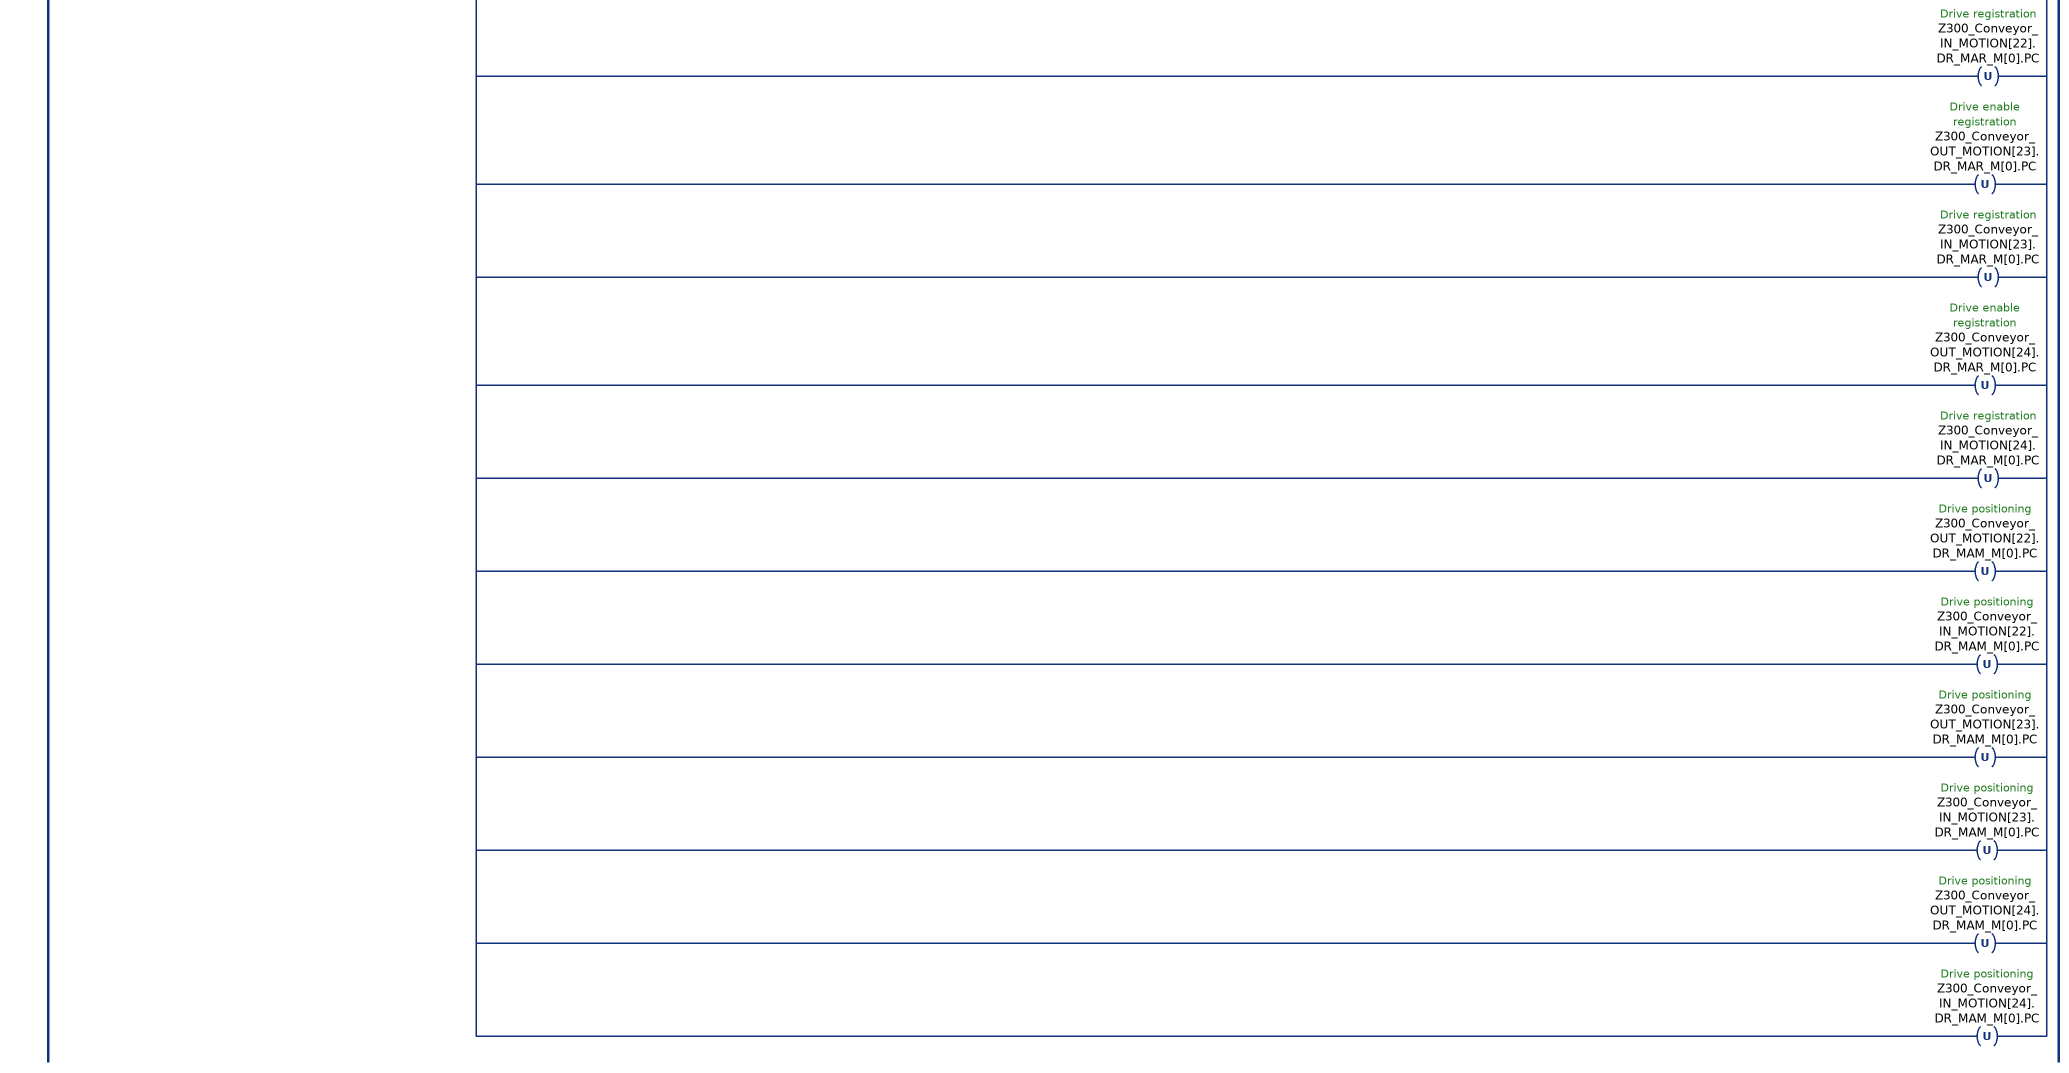
   // Positioning request (In case of head positioning also previous conveyors are involved)
   32: XIO(M310Popup[0].ST_xPlateInPositionToRise)XIO(M310Popup[1].ST_xPlateInPositionToRise)XIC(M310Popup[0].AUX_tSearchPlateData.xPlateHooked)[XIC(M310Popup[0].ST_xPlateToSinglePositioning) XIO(Z300_LineTracking.rgtTrkConv[22].xGlassPresence) XIO(Z300_LineTracking.rgtTrkConv[23].xGlassPresence) XIO(M310Popup[0].ST_xPlatePresence) [XIO(M310Popup[0].ST_xPlateUnderPopup) ,XIO(xDebugOFF) ] XIC(M310Popup[0].ST_xOutputEnable) XIC(M310Popup[0].INPUT_xPopupLow) XIC(M310Popup[0].ST_xInitialConditionForRise) ,XIC(M310Popup[1].ST_xPlateToSinglePositioning) XIO(Z300_LineTracking.rgtTrkConv[22].xGlassPresence) XIO(Z300_LineTracking.rgtTrkConv[23].xGlassPresence) XIO(Z300_LineTracking.rgtTrkConv[24].xGlassPresence) XIO(M310Popup[1].ST_xPlatePresence) XIO(M310Popup[0].ST_xPlateUnderPopup) [XIO(M310Popup[1].ST_xPlateUnderPopup) ,XIO(xDebugOFF) ] XIC(M310Popup[1].ST_xOutputEnable) XIC(M310Popup[1].INPUT_xPopupLow) XIC(M310Popup[1].ST_xInitialConditionForRise) ,XIC(M310Popup[0].ST_xPlateToBothPositioning) XIO(Z300_LineTracking.rgtTrkConv[22].xGlassPresence) XIO(Z300_LineTracking.rgtTrkConv[23].xGlassPresence) XIO(Z300_LineTracking.rgtTrkConv[24].xGlassPresence) XIO(M310Popup[0].ST_xPlatePresence) XIO(M310Popup[0].ST_xPlateUnderPopup) XIC(M310Popup[0].ST_xOutputEnable) XIC(M310Popup[0].INPUT_xPopupLow) XIC(M310Popup[0].ST_xInitialConditionForRise) XIO(M310Popup[1].ST_xPlatePresence) [XIO(M310Popup[1].ST_xPlateUnderPopup) ,XIO(xDebugOFF) ] XIC(M310Popup[1].ST_xOutputEnable) XIC(M310Popup[1].INPUT_xPopupLow) XIC(M310Popup[1].ST_xInitialConditionForRise) ,XIC(M310Popup[0].ST_xConvoyPositioning) XIO(Z300_LineTracking.rgtTrkConv[22].xGlassPresence) XIO(Z300_LineTracking.rgtTrkConv[23].xGlassPresence) XIO(Z300_LineTracking.rgtTrkConv[24].xGlassPresence) XIO(M310Popup[0].ST_xPlatePresence) XIO(M310Popup[0].ST_xPlateUnderPopup) XIC(M310Popup[0].ST_xOutputEnable) XIC(M310Popup[0].INPUT_xPopupLow) XIC(M310Popup[0].ST_xInitialConditionForRise) XIO(M310Popup[1].ST_xPlatePresence) [XIO(M310Popup[1].ST_xPlateUnderPopup) ,XIO(xDebugOFF) ] XIC(M310Popup[1].ST_xOutputEnable) XIC(M310Popup[1].INPUT_xPopupLow) XIC(M310Popup[1].ST_xInitialConditionForRise) ]XIO(Z300_Conveyor[22].xReqStop)XIO(Z300_Conveyor[23].xReqStop)[XIC(M310Popup[0].ST_xIndexConsPositioning) ,XIO(xDebugOFF) ][XIC(TMP_xPosHead) XIC(M310Popup[0].AUX_tSearchPlateData.tResult.xHeadPresence) ,XIO(TMP_xPosHead) XIC(M310Popup[0].AUX_tSearchPlateData.tResult.xTailPresence) ]XIO(Z300_Conveyor[22].xReqPositioningHead)XIO(Z300_Conveyor[22].xReqPositioningTail)XIO(Z300_Conveyor[23].xReqPositioningHead)XIO(Z300_Conveyor[23].xReqPositioningTail)[XIO(Z300_Conveyor[24].xReqStop) XIO(Z300_Conveyor[24].xReqPositioningHead) XIO(Z300_Conveyor[24].xReqPositioningTail) ,XIC(M310Popup[1].ST_xPlateToSinglePositioning) ]XIO(M310Popup[0].tmOF_Wait.DN)XIO(M310Popup[1].tmOF_Wait.DN)TON(M310Popup[0].tmON_Positioning,?,?)XIC(M310Popup[0].tmON_Positioning.DN)[XIC(TMP_xPosHead) [OTL(Z300_Conveyor[22].xReqPositioningHead) ,OTL(Z300_Conveyor[23].xReqPositioningHead) ] ,XIO(TMP_xPosHead) [OTL(Z300_Conveyor[22].xReqPositioningTail) ,OTL(Z300_Conveyor[23].xReqPositioningTail) ] ,OTE(M310Popup[0].OS_xStartPositioning) ,[XIC(M310Popup[0].ST_xPlateToBothPositioning) ,XIC(M310Popup[0].ST_xConvoyPositioning) ,XIC(M310Popup[1].ST_xPlateToSinglePositioning) ] [XIC(TMP_xPosHead) OTL(Z300_Conveyor[24].xReqPositioningHead) ,XIO(TMP_xPosHead) OTL(Z300_Conveyor[24].xReqPositioningTail) ,OTE(M310Popup[1].OS_xStartPositioning) ] ,OTU(Z300_Conveyor_OUT_MOTION[22].DR_MAR_M[0].PC) ,OTU(Z300_Conveyor_IN_MOTION[22].DR_MAR_M[0].PC) ,OTU(Z300_Conveyor_OUT_MOTION[23].DR_MAR_M[0].PC) ,OTU(Z300_Conveyor_IN_MOTION[23].DR_MAR_M[0].PC) ,OTU(Z300_Conveyor_OUT_MOTION[24].DR_MAR_M[0].PC) ,OTU(Z300_Conveyor_IN_MOTION[24].DR_MAR_M[0].PC) ,OTU(Z300_Conveyor_OUT_MOTION[22].DR_MAM_M[0].PC) ,OTU(Z300_Conveyor_IN_MOTION[22].DR_MAM_M[0].PC) ,OTU(Z300_Conveyor_OUT_MOTION[23].DR_MAM_M[0].PC) ,OTU(Z300_Conveyor_IN_MOTION[23].DR_MAM_M[0].PC) ,OTU(Z300_Conveyor_OUT_MOTION[24].DR_MAM_M[0].PC) ,OTU(Z300_Conveyor_IN_MOTION[24].DR_MAM_M[0].PC) ];
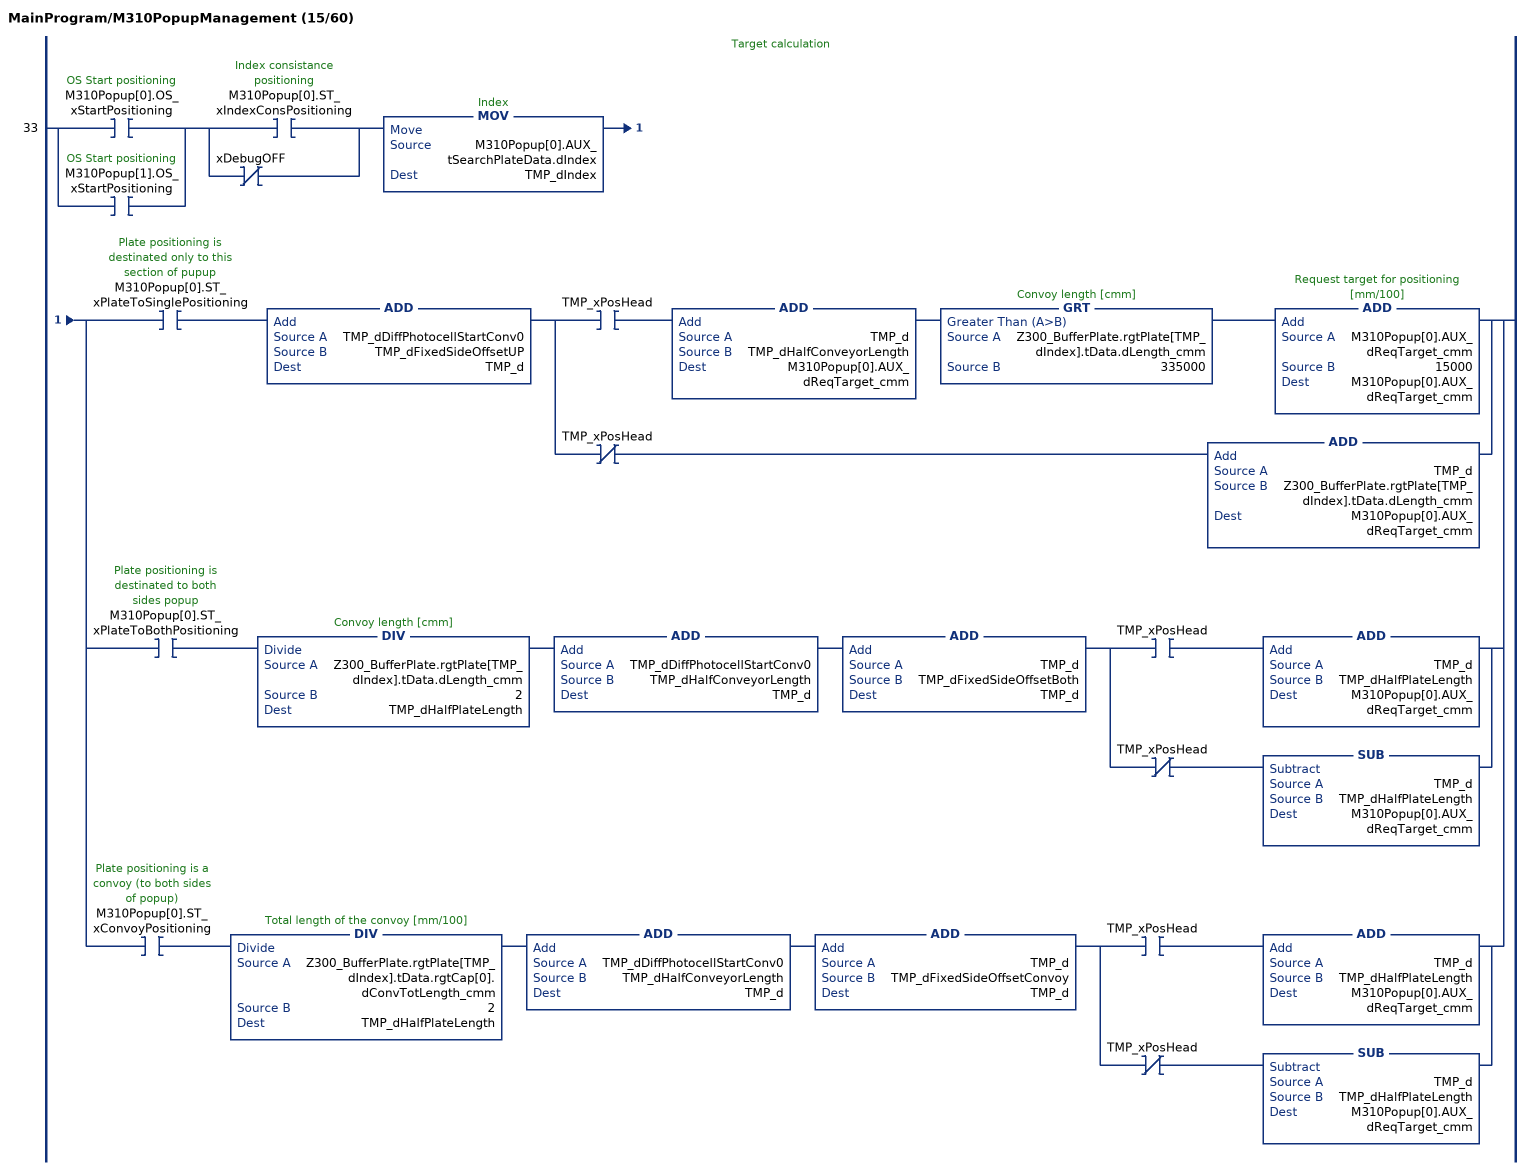
   // Target calculation
   33: [XIC(M310Popup[0].OS_xStartPositioning) ,XIC(M310Popup[1].OS_xStartPositioning) ][XIC(M310Popup[0].ST_xIndexConsPositioning) ,XIO(xDebugOFF) ]MOV(M310Popup[0].AUX_tSearchPlateData.dIndex,TMP_dIndex)[XIC(M310Popup[0].ST_xPlateToSinglePositioning) ADD(TMP_dDiffPhotocellStartConv0,TMP_dFixedSideOffsetUP,TMP_d) [XIC(TMP_xPosHead) ADD(TMP_d,TMP_dHalfConveyorLength,M310Popup[0].AUX_dReqTarget_cmm) GRT(Z300_BufferPlate.rgtPlate[TMP_dIndex].tData.dLength_cmm,335000) ADD(M310Popup[0].AUX_dReqTarget_cmm,15000,M310Popup[0].AUX_dReqTarget_cmm) ,XIO(TMP_xPosHead) ADD(TMP_d,Z300_BufferPlate.rgtPlate[TMP_dIndex].tData.dLength_cmm,M310Popup[0].AUX_dReqTarget_cmm) ] ,XIC(M310Popup[0].ST_xPlateToBothPositioning) DIV(Z300_BufferPlate.rgtPlate[TMP_dIndex].tData.dLength_cmm,2,TMP_dHalfPlateLength) ADD(TMP_dDiffPhotocellStartConv0,TMP_dHalfConveyorLength,TMP_d) ADD(TMP_d,TMP_dFixedSideOffsetBoth,TMP_d) [XIC(TMP_xPosHead) ADD(TMP_d,TMP_dHalfPlateLength,M310Popup[0].AUX_dReqTarget_cmm) ,XIO(TMP_xPosHead) SUB(TMP_d,TMP_dHalfPlateLength,M310Popup[0].AUX_dReqTarget_cmm) ] ,XIC(M310Popup[0].ST_xConvoyPositioning) DIV(Z300_BufferPlate.rgtPlate[TMP_dIndex].tData.rgtCap[0].dConvTotLength_cmm,2,TMP_dHalfPlateLength) ADD(TMP_dDiffPhotocellStartConv0,TMP_dHalfConveyorLength,TMP_d) ADD(TMP_d,TMP_dFixedSideOffsetConvoy,TMP_d) [XIC(TMP_xPosHead) ADD(TMP_d,TMP_dHalfPlateLength,M310Popup[0].AUX_dReqTarget_cmm) ,XIO(TMP_xPosHead) SUB(TMP_d,TMP_dHalfPlateLength,M310Popup[0].AUX_dReqTarget_cmm) ] ];
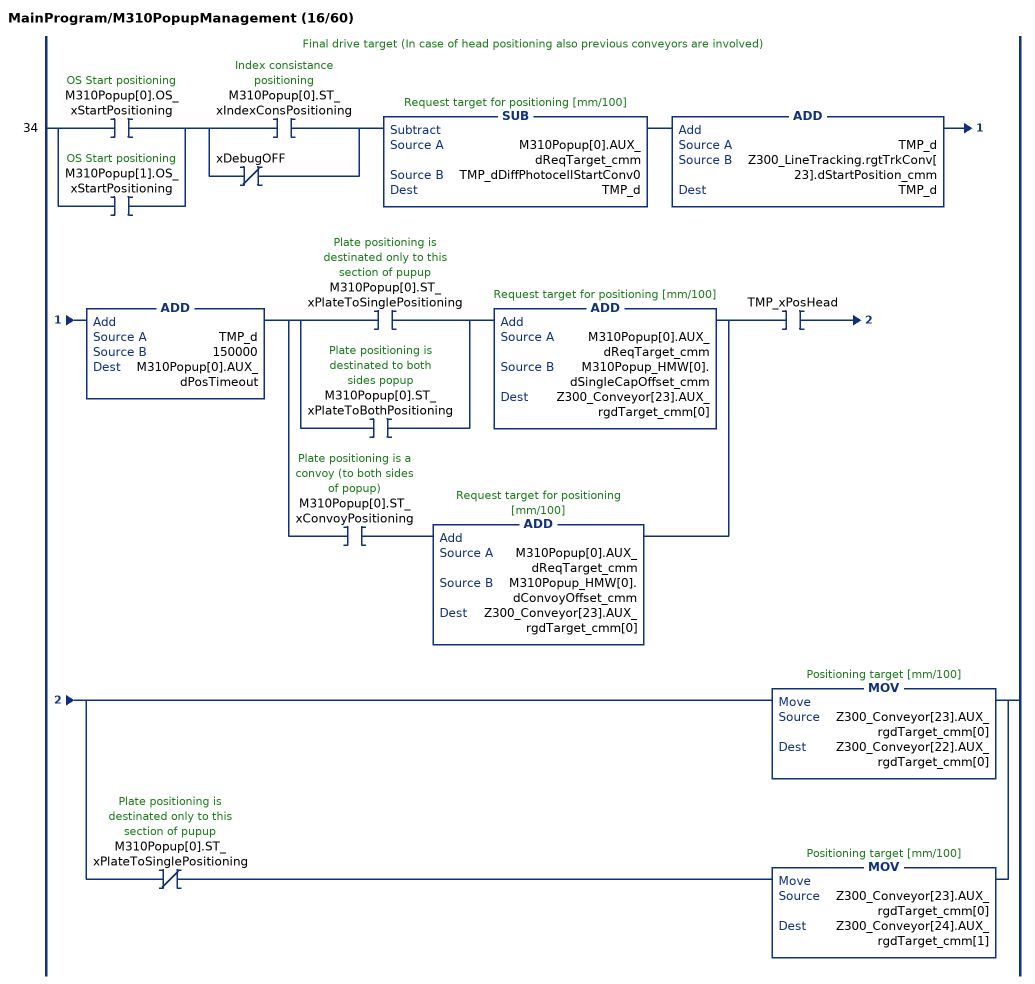
   // Final drive target (In case of head positioning also previous conveyors are involved)
   34: [XIC(M310Popup[0].OS_xStartPositioning) ,XIC(M310Popup[1].OS_xStartPositioning) ][XIC(M310Popup[0].ST_xIndexConsPositioning) ,XIO(xDebugOFF) ]SUB(M310Popup[0].AUX_dReqTarget_cmm,TMP_dDiffPhotocellStartConv0,TMP_d)ADD(TMP_d,Z300_LineTracking.rgtTrkConv[23].dStartPosition_cmm,TMP_d)ADD(TMP_d,150000,M310Popup[0].AUX_dPosTimeout)[[XIC(M310Popup[0].ST_xPlateToSinglePositioning) ,XIC(M310Popup[0].ST_xPlateToBothPositioning) ] ADD(M310Popup[0].AUX_dReqTarget_cmm,M310Popup_HMW[0].dSingleCapOffset_cmm,Z300_Conveyor[23].AUX_rgdTarget_cmm[0]) ,XIC(M310Popup[0].ST_xConvoyPositioning) ADD(M310Popup[0].AUX_dReqTarget_cmm,M310Popup_HMW[0].dConvoyOffset_cmm,Z300_Conveyor[23].AUX_rgdTarget_cmm[0]) ]XIC(TMP_xPosHead)[MOV(Z300_Conveyor[23].AUX_rgdTarget_cmm[0],Z300_Conveyor[22].AUX_rgdTarget_cmm[0]) ,XIO(M310Popup[0].ST_xPlateToSinglePositioning) MOV(Z300_Conveyor[23].AUX_rgdTarget_cmm[0],Z300_Conveyor[24].AUX_rgdTarget_cmm[1]) ];
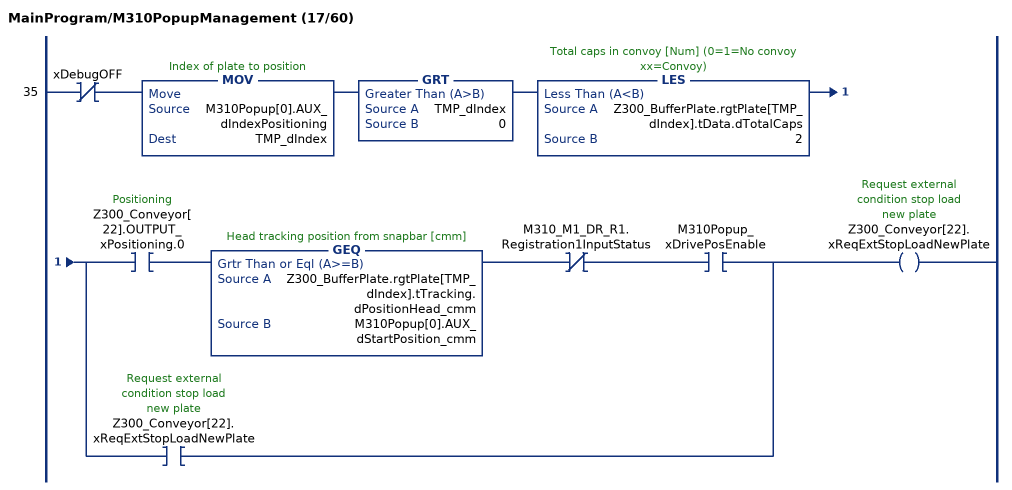
   35: XIO(xDebugOFF)MOV(M310Popup[0].AUX_dIndexPositioning,TMP_dIndex)GRT(TMP_dIndex,0)LES(Z300_BufferPlate.rgtPlate[TMP_dIndex].tData.dTotalCaps,2)[XIC(Z300_Conveyor[22].OUTPUT_xPositioning.0) GEQ(Z300_BufferPlate.rgtPlate[TMP_dIndex].tTracking.dPositionHead_cmm,M310Popup[0].AUX_dStartPosition_cmm) XIO(M310_M1_DR_R1.Registration1InputStatus) XIC(M310Popup_xDrivePosEnable) ,XIC(Z300_Conveyor[22].xReqExtStopLoadNewPlate) ]OTE(Z300_Conveyor[22].xReqExtStopLoadNewPlate);
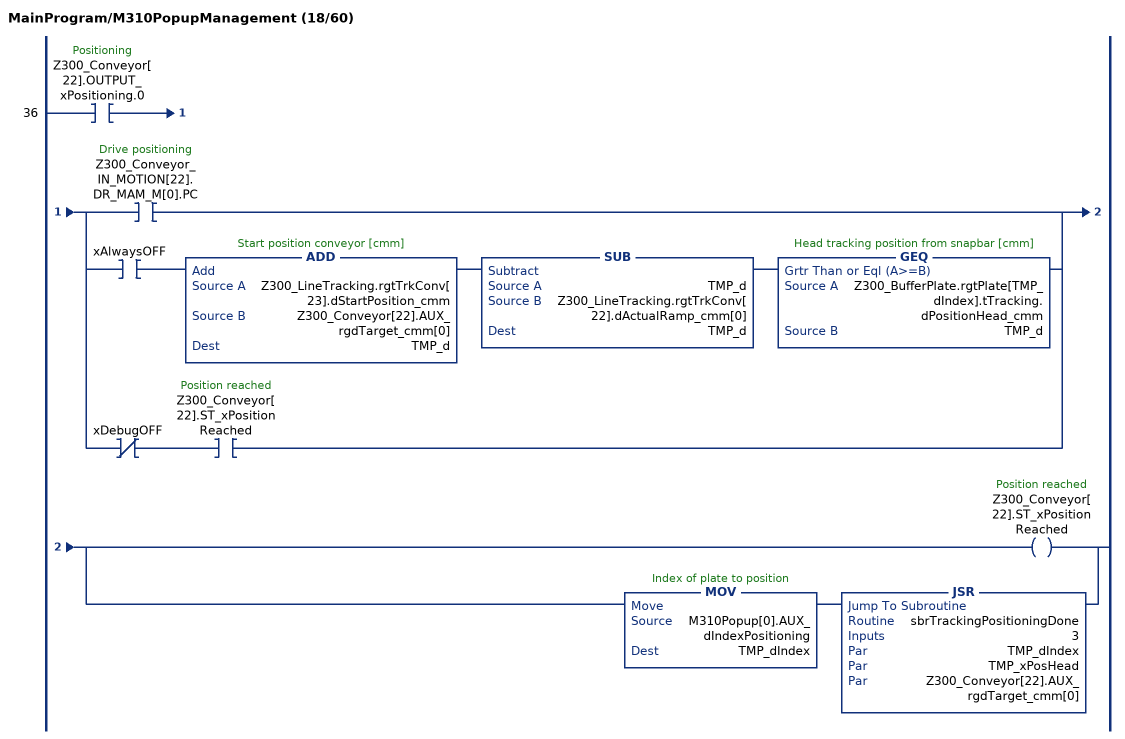
   36: XIC(Z300_Conveyor[22].OUTPUT_xPositioning.0)[[XIC(Z300_Conveyor_IN_MOTION[22].DR_MAM_M[0].PC) ,XIC(xAlwaysOFF) ADD(Z300_LineTracking.rgtTrkConv[23].dStartPosition_cmm,Z300_Conveyor[22].AUX_rgdTarget_cmm[0],TMP_d) SUB(TMP_d,Z300_LineTracking.rgtTrkConv[22].dActualRamp_cmm[0],TMP_d) GEQ(Z300_BufferPlate.rgtPlate[TMP_dIndex].tTracking.dPositionHead_cmm,TMP_d) ] ,XIO(xDebugOFF) XIC(Z300_Conveyor[22].ST_xPositionReached) ][OTE(Z300_Conveyor[22].ST_xPositionReached) ,MOV(M310Popup[0].AUX_dIndexPositioning,TMP_dIndex) JSR(sbrTrackingPositioningDone,3,TMP_dIndex,TMP_xPosHead,Z300_Conveyor[22].AUX_rgdTarget_cmm[0]) ];
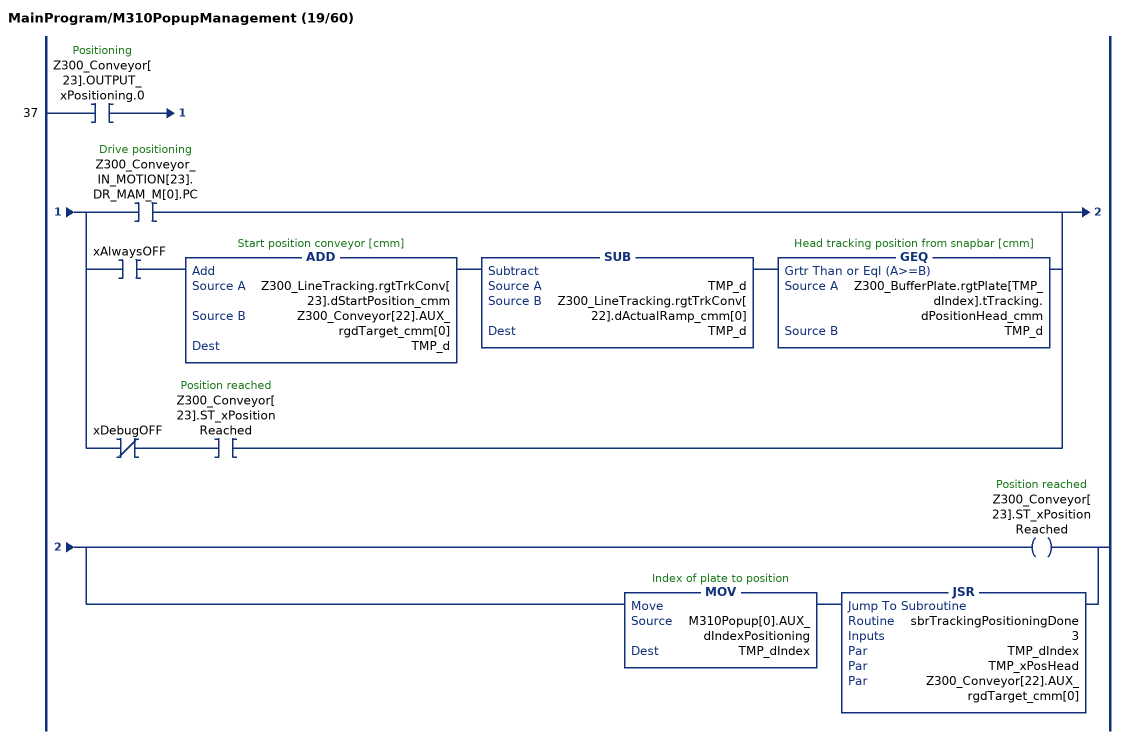
   37: XIC(Z300_Conveyor[23].OUTPUT_xPositioning.0)[[XIC(Z300_Conveyor_IN_MOTION[23].DR_MAM_M[0].PC) ,XIC(xAlwaysOFF) ADD(Z300_LineTracking.rgtTrkConv[23].dStartPosition_cmm,Z300_Conveyor[22].AUX_rgdTarget_cmm[0],TMP_d) SUB(TMP_d,Z300_LineTracking.rgtTrkConv[22].dActualRamp_cmm[0],TMP_d) GEQ(Z300_BufferPlate.rgtPlate[TMP_dIndex].tTracking.dPositionHead_cmm,TMP_d) ] ,XIO(xDebugOFF) XIC(Z300_Conveyor[23].ST_xPositionReached) ][OTE(Z300_Conveyor[23].ST_xPositionReached) ,MOV(M310Popup[0].AUX_dIndexPositioning,TMP_dIndex) JSR(sbrTrackingPositioningDone,3,TMP_dIndex,TMP_xPosHead,Z300_Conveyor[22].AUX_rgdTarget_cmm[0]) ];
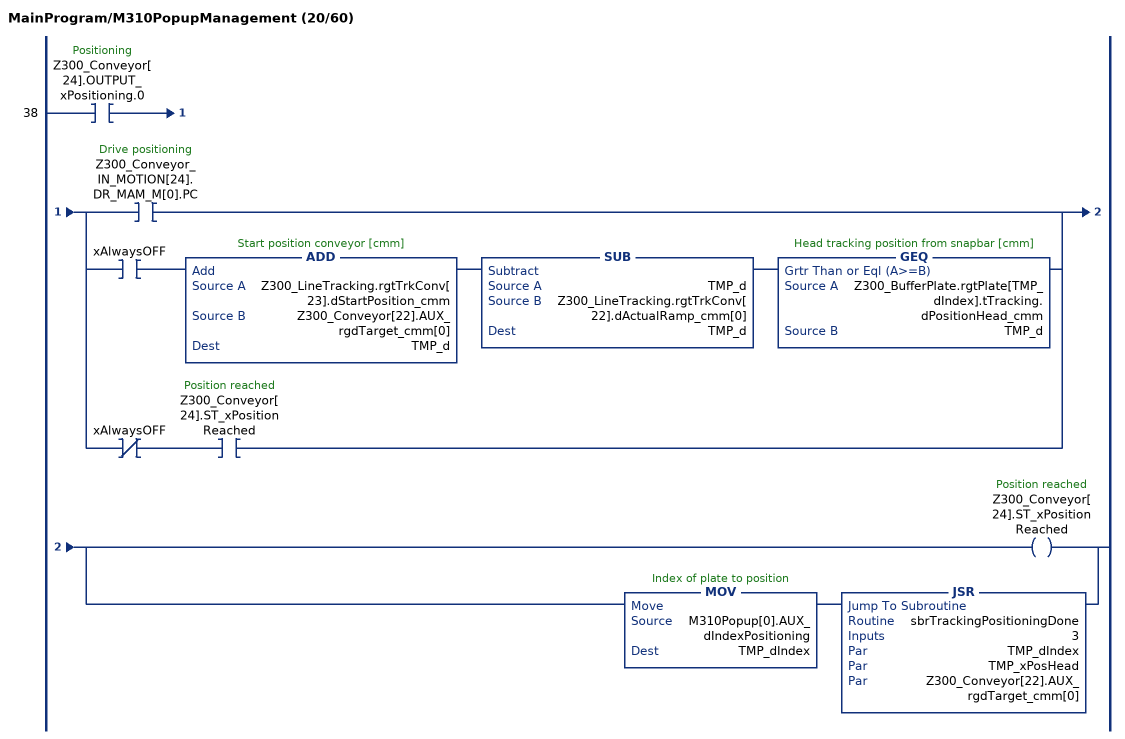
   38: XIC(Z300_Conveyor[24].OUTPUT_xPositioning.0)[XIC(Z300_Conveyor_IN_MOTION[24].DR_MAM_M[0].PC) ,XIC(xAlwaysOFF) ADD(Z300_LineTracking.rgtTrkConv[23].dStartPosition_cmm,Z300_Conveyor[22].AUX_rgdTarget_cmm[0],TMP_d) SUB(TMP_d,Z300_LineTracking.rgtTrkConv[22].dActualRamp_cmm[0],TMP_d) GEQ(Z300_BufferPlate.rgtPlate[TMP_dIndex].tTracking.dPositionHead_cmm,TMP_d) ,XIO(xAlwaysOFF) XIC(Z300_Conveyor[24].ST_xPositionReached) ][OTE(Z300_Conveyor[24].ST_xPositionReached) ,MOV(M310Popup[0].AUX_dIndexPositioning,TMP_dIndex) JSR(sbrTrackingPositioningDone,3,TMP_dIndex,TMP_xPosHead,Z300_Conveyor[22].AUX_rgdTarget_cmm[0]) ];
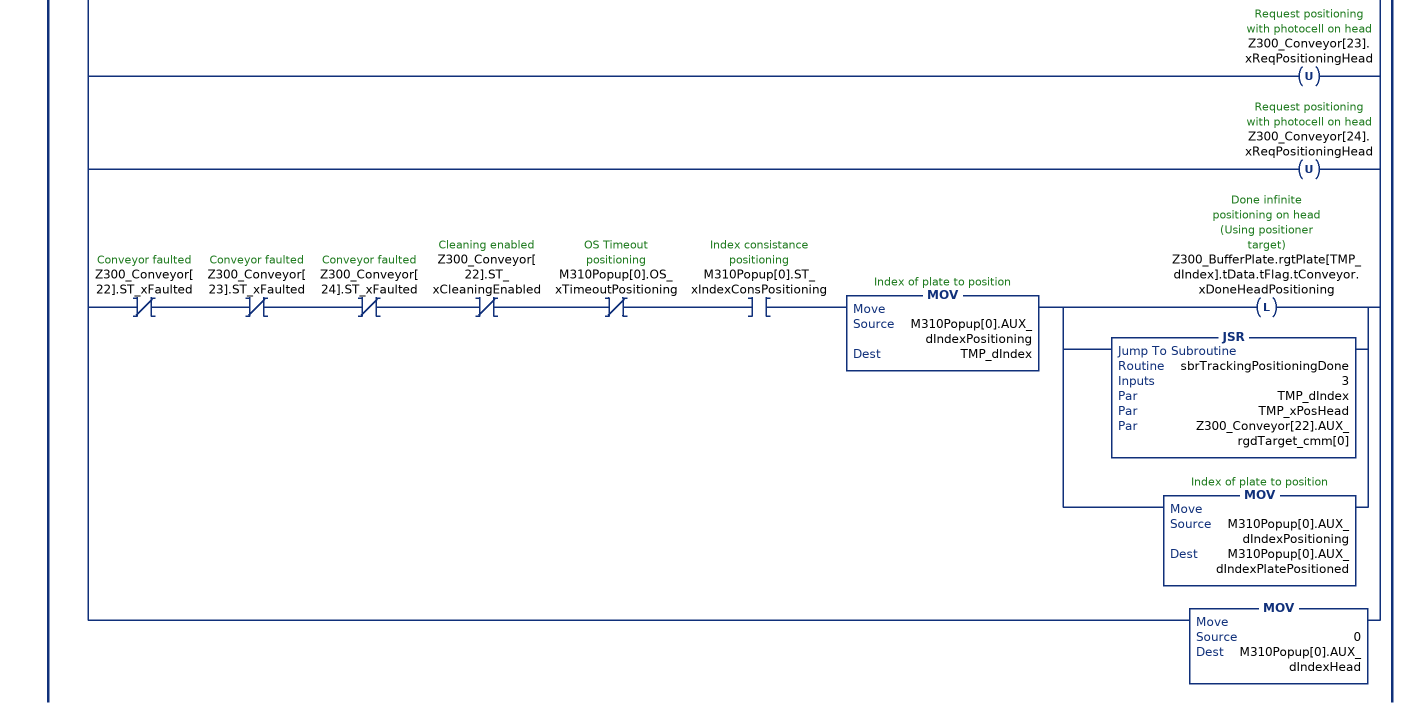
   // Head positioning done
   39: [XIC(Z300_Conveyor[22].xReqPositioningHead) ,XIC(Z300_Conveyor[23].xReqPositioningHead) ,XIC(Z300_Conveyor[24].xReqPositioningHead) ][XIC(Z300_Conveyor[22].ST_xPositionReached) XIC(Z300_Conveyor[23].ST_xPositionReached) [XIC(Z300_Conveyor[24].ST_xPositionReached) ,XIO(Z300_Conveyor[24].xReqPositioningHead) ] ,XIC(Z300_Conveyor[22].xReqStop) XIO(Z300_Conveyor[22].ST_xRotationFeedback) XIC(Z300_Conveyor[23].xReqStop) XIO(Z300_Conveyor[23].ST_xRotationFeedback) [XIC(Z300_Conveyor[24].xReqStop) XIO(Z300_Conveyor[24].ST_xRotationFeedback) ,XIO(Z300_Conveyor[24].xReqPositioningHead) ] ,XIC(M310Popup[0].OS_xTimeoutPositioning) ,XIC(xDebugOFF) XIO(M310Popup[0].ST_xIndexConsPositioning) ,XIC(Z300_Conveyor[23].ST_xCleaningEnabled) ,XIC(Z300_Conveyor[22].ST_xFaulted) ,XIC(Z300_Conveyor[23].ST_xFaulted) ,XIC(Z300_Conveyor[24].ST_xFaulted) ][OTU(Z300_Conveyor[22].xReqPositioningHead) ,OTU(Z300_Conveyor[23].xReqPositioningHead) ,OTU(Z300_Conveyor[24].xReqPositioningHead) ,XIO(Z300_Conveyor[22].ST_xFaulted) XIO(Z300_Conveyor[23].ST_xFaulted) XIO(Z300_Conveyor[24].ST_xFaulted) XIO(Z300_Conveyor[22].ST_xCleaningEnabled) XIO(M310Popup[0].OS_xTimeoutPositioning) XIC(M310Popup[0].ST_xIndexConsPositioning) MOV(M310Popup[0].AUX_dIndexPositioning,TMP_dIndex) [OTL(Z300_BufferPlate.rgtPlate[TMP_dIndex].tData.tFlag.tConveyor.xDoneHeadPositioning) ,JSR(sbrTrackingPositioningDone,3,TMP_dIndex,TMP_xPosHead,Z300_Conveyor[22].AUX_rgdTarget_cmm[0]) ,MOV(M310Popup[0].AUX_dIndexPositioning,M310Popup[0].AUX_dIndexPlatePositioned) ] ,MOV(0,M310Popup[0].AUX_dIndexHead) ];
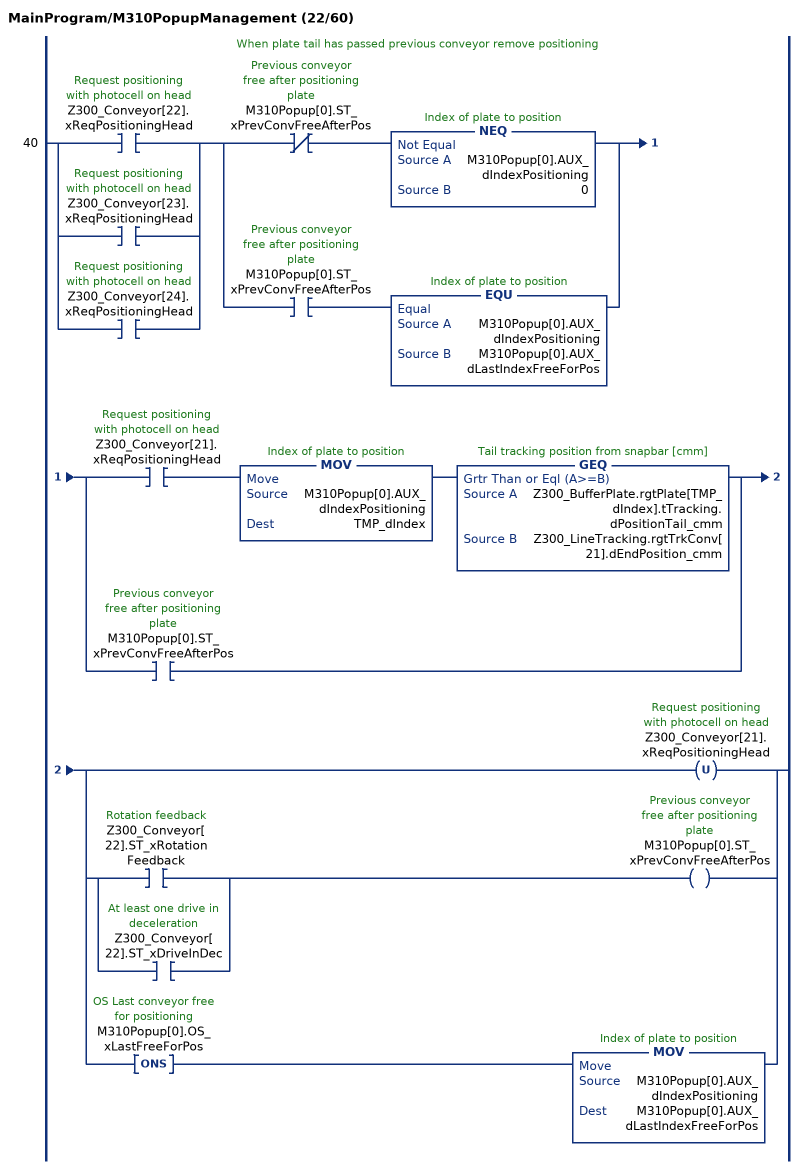
   // When plate tail has passed previous conveyor remove positioning
   40: [XIC(Z300_Conveyor[22].xReqPositioningHead) ,XIC(Z300_Conveyor[23].xReqPositioningHead) ,XIC(Z300_Conveyor[24].xReqPositioningHead) ][XIO(M310Popup[0].ST_xPrevConvFreeAfterPos) NEQ(M310Popup[0].AUX_dIndexPositioning,0) ,XIC(M310Popup[0].ST_xPrevConvFreeAfterPos) EQU(M310Popup[0].AUX_dIndexPositioning,M310Popup[0].AUX_dLastIndexFreeForPos) ][XIC(Z300_Conveyor[21].xReqPositioningHead) MOV(M310Popup[0].AUX_dIndexPositioning,TMP_dIndex) GEQ(Z300_BufferPlate.rgtPlate[TMP_dIndex].tTracking.dPositionTail_cmm,Z300_LineTracking.rgtTrkConv[21].dEndPosition_cmm) ,XIC(M310Popup[0].ST_xPrevConvFreeAfterPos) ][OTU(Z300_Conveyor[21].xReqPositioningHead) ,[XIC(Z300_Conveyor[22].ST_xRotationFeedback) ,XIC(Z300_Conveyor[22].ST_xDriveInDec) ] OTE(M310Popup[0].ST_xPrevConvFreeAfterPos) ,ONS(M310Popup[0].OS_xLastFreeForPos) MOV(M310Popup[0].AUX_dIndexPositioning,M310Popup[0].AUX_dLastIndexFreeForPos) ];
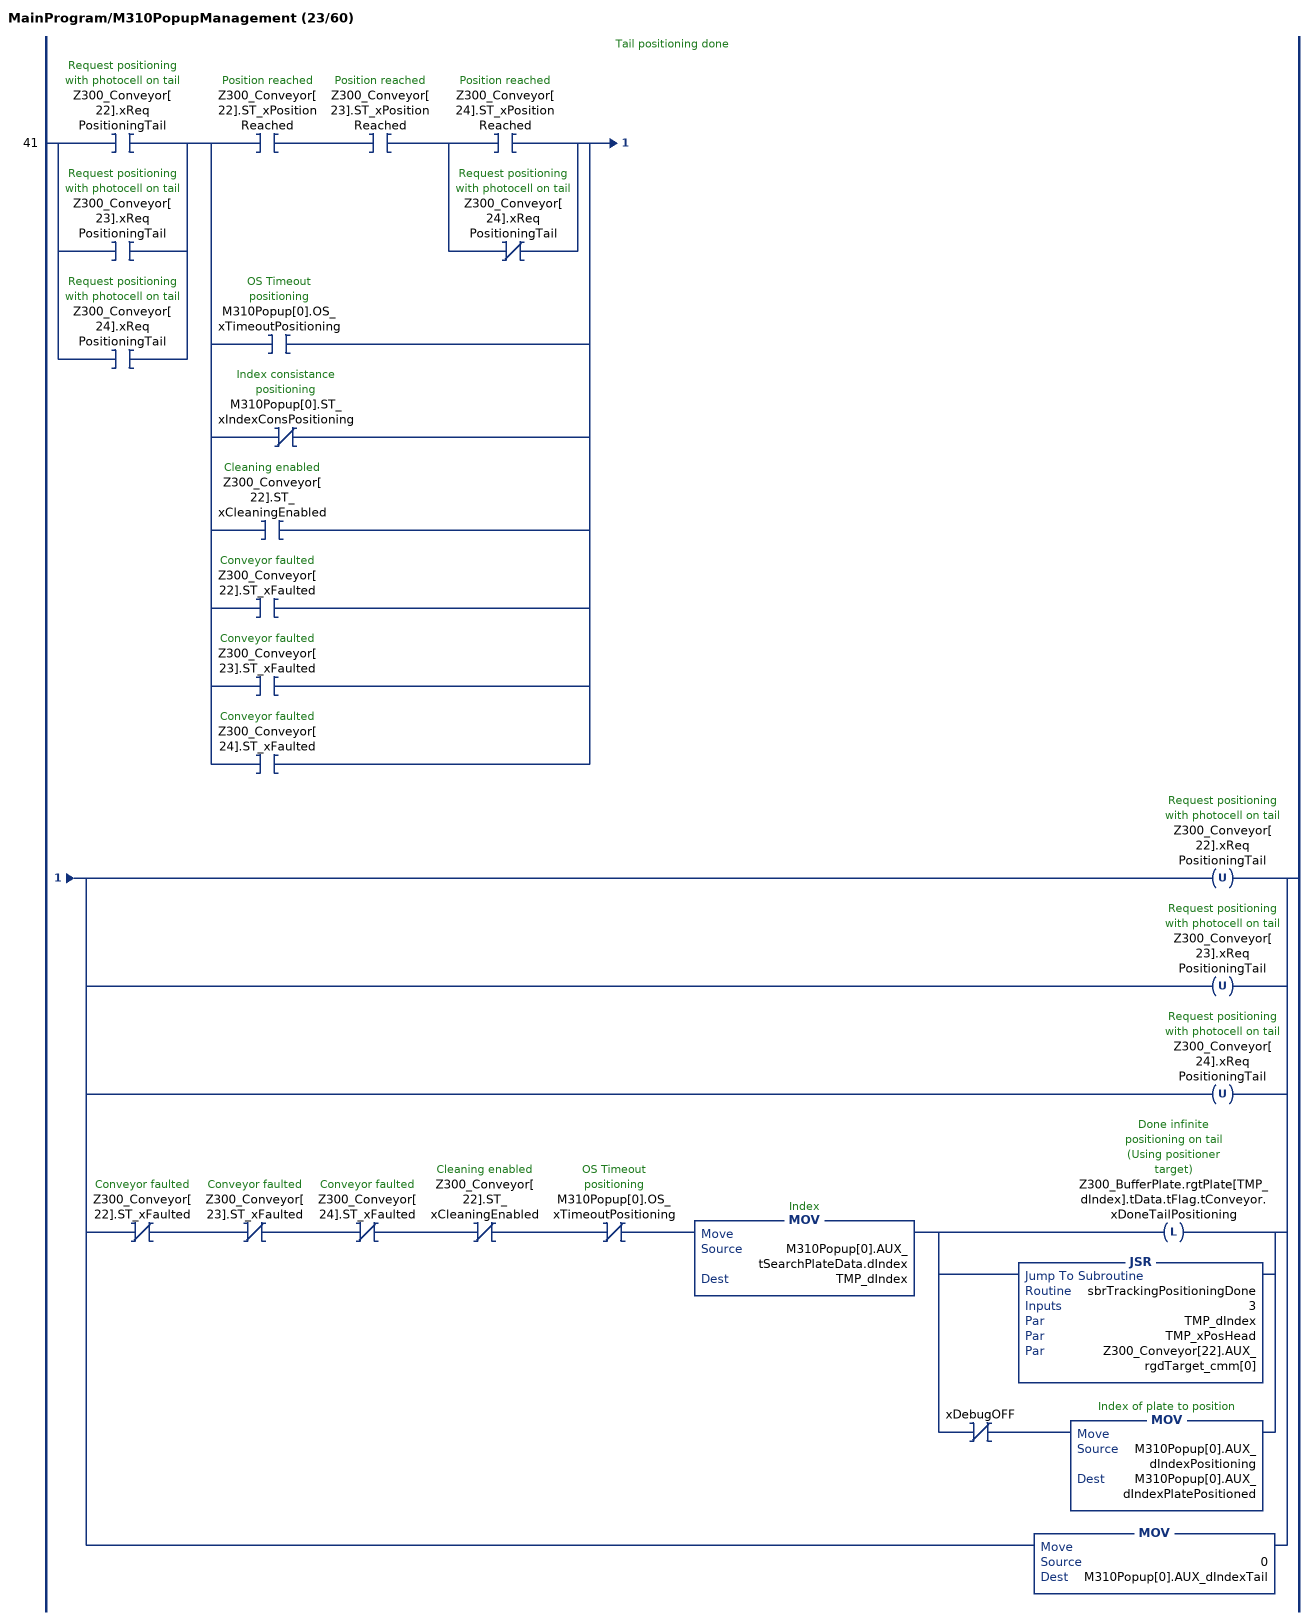
   // Tail positioning done
   41: [XIC(Z300_Conveyor[22].xReqPositioningTail) ,XIC(Z300_Conveyor[23].xReqPositioningTail) ,XIC(Z300_Conveyor[24].xReqPositioningTail) ][XIC(Z300_Conveyor[22].ST_xPositionReached) XIC(Z300_Conveyor[23].ST_xPositionReached) [XIC(Z300_Conveyor[24].ST_xPositionReached) ,XIO(Z300_Conveyor[24].xReqPositioningTail) ] ,XIC(M310Popup[0].OS_xTimeoutPositioning) ,XIO(M310Popup[0].ST_xIndexConsPositioning) ,XIC(Z300_Conveyor[22].ST_xCleaningEnabled) ,XIC(Z300_Conveyor[22].ST_xFaulted) ,XIC(Z300_Conveyor[23].ST_xFaulted) ,XIC(Z300_Conveyor[24].ST_xFaulted) ][OTU(Z300_Conveyor[22].xReqPositioningTail) ,OTU(Z300_Conveyor[23].xReqPositioningTail) ,OTU(Z300_Conveyor[24].xReqPositioningTail) ,XIO(Z300_Conveyor[22].ST_xFaulted) XIO(Z300_Conveyor[23].ST_xFaulted) XIO(Z300_Conveyor[24].ST_xFaulted) XIO(Z300_Conveyor[22].ST_xCleaningEnabled) XIO(M310Popup[0].OS_xTimeoutPositioning) MOV(M310Popup[0].AUX_tSearchPlateData.dIndex,TMP_dIndex) [OTL(Z300_BufferPlate.rgtPlate[TMP_dIndex].tData.tFlag.tConveyor.xDoneTailPositioning) ,JSR(sbrTrackingPositioningDone,3,TMP_dIndex,TMP_xPosHead,Z300_Conveyor[22].AUX_rgdTarget_cmm[0]) ,XIO(xDebugOFF) MOV(M310Popup[0].AUX_dIndexPositioning,M310Popup[0].AUX_dIndexPlatePositioned) ] ,MOV(0,M310Popup[0].AUX_dIndexTail) ];
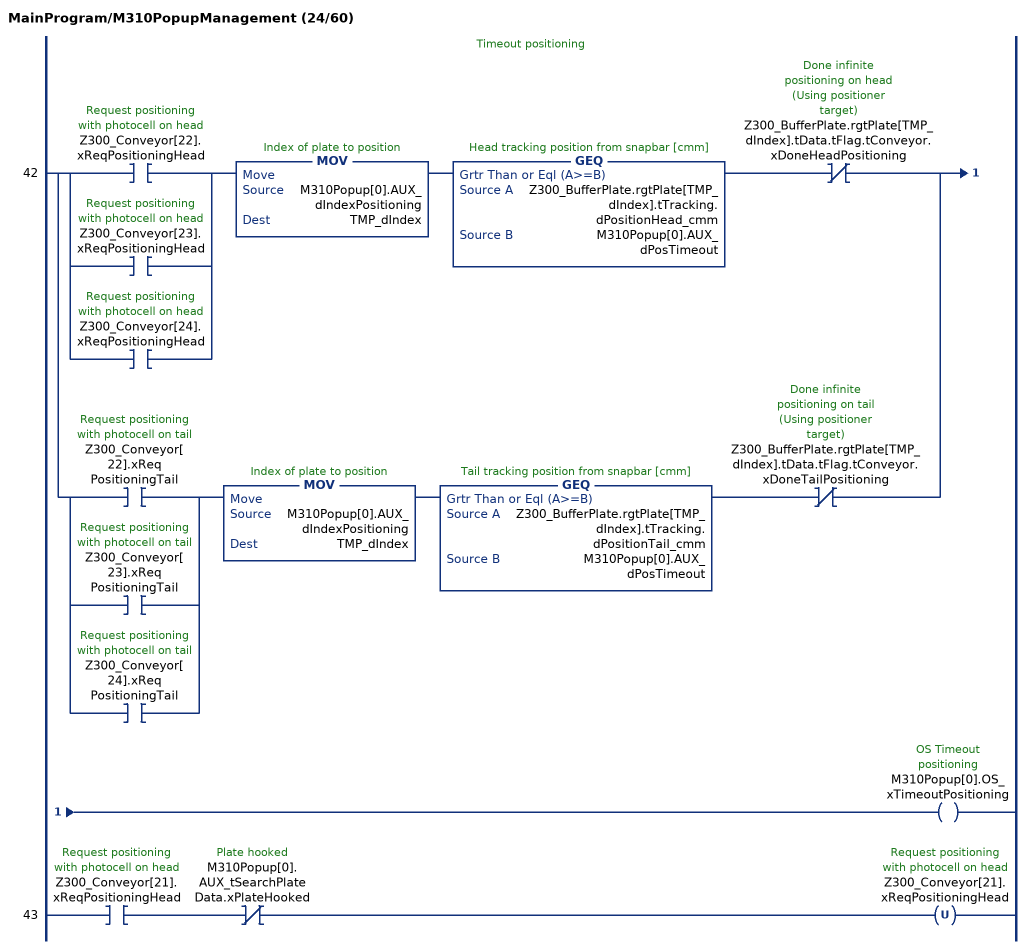
   // Timeout positioning
   42: [[XIC(Z300_Conveyor[22].xReqPositioningHead) ,XIC(Z300_Conveyor[23].xReqPositioningHead) ,XIC(Z300_Conveyor[24].xReqPositioningHead) ] MOV(M310Popup[0].AUX_dIndexPositioning,TMP_dIndex) GEQ(Z300_BufferPlate.rgtPlate[TMP_dIndex].tTracking.dPositionHead_cmm,M310Popup[0].AUX_dPosTimeout) XIO(Z300_BufferPlate.rgtPlate[TMP_dIndex].tData.tFlag.tConveyor.xDoneHeadPositioning) ,[XIC(Z300_Conveyor[22].xReqPositioningTail) ,XIC(Z300_Conveyor[23].xReqPositioningTail) ,XIC(Z300_Conveyor[24].xReqPositioningTail) ] MOV(M310Popup[0].AUX_dIndexPositioning,TMP_dIndex) GEQ(Z300_BufferPlate.rgtPlate[TMP_dIndex].tTracking.dPositionTail_cmm,M310Popup[0].AUX_dPosTimeout) XIO(Z300_BufferPlate.rgtPlate[TMP_dIndex].tData.tFlag.tConveyor.xDoneTailPositioning) ]OTE(M310Popup[0].OS_xTimeoutPositioning);
   43: XIC(Z300_Conveyor[21].xReqPositioningHead)XIO(M310Popup[0].AUX_tSearchPlateData.xPlateHooked)OTU(Z300_Conveyor[21].xReqPositioningHead);
